REGION Network 10: Ethernet.Enc2 Too big speed change
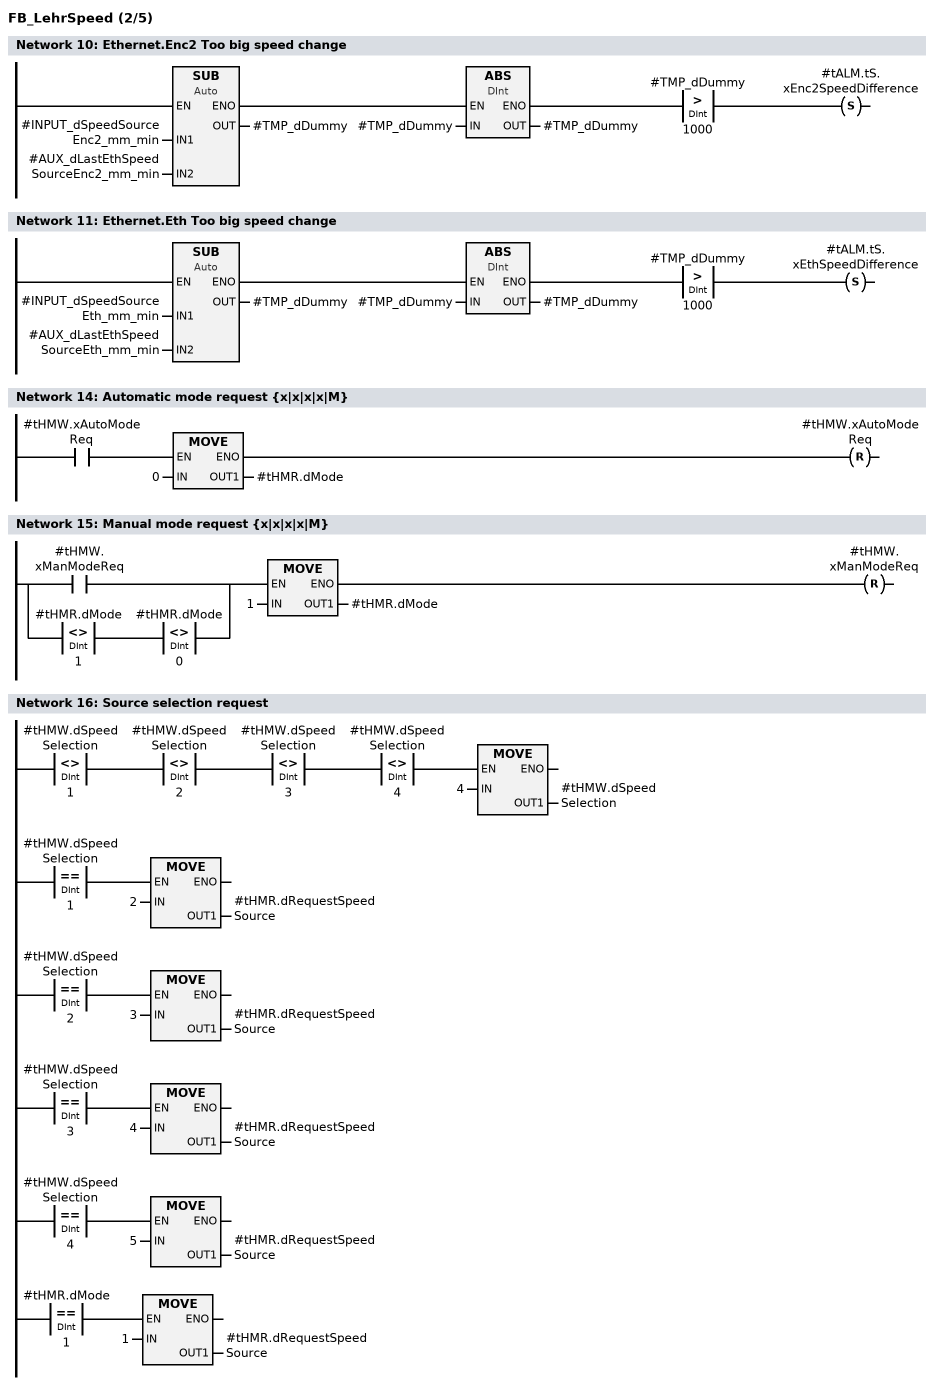
   RUNG wire#powerrail
      Sub(in1 := #INPUT_dSpeedSourceEnc2_mm_min, in2 := #AUX_dLastEthSpeedSourceEnc2_mm_min, out => #TMP_dDummy)
      { S7_Templates := "SrcType := DInt" } Abs(in := #TMP_dDummy, out => #TMP_dDummy)
      { S7_Templates := "SrcType := DInt" } GT_Contact(in1 := #TMP_dDummy, in2 := 1000)
      S_Coil( #tALM.tS.xEnc2SpeedDifference )
   END_RUNG
   // the same network as SCL:
   #TMP_dDummy := #INPUT_dSpeedSourceEnc2_mm_min - #AUX_dLastEthSpeedSourceEnc2_mm_min;
   #TMP_dDummy := ABS(#TMP_dDummy);
   IF #TMP_dDummy > 1000 THEN #tALM.tS.xEnc2SpeedDifference := TRUE; END_IF;
END_REGION

REGION Network 11: Ethernet.Eth Too big speed change
   RUNG wire#powerrail
      Sub(in1 := #INPUT_dSpeedSourceEth_mm_min, in2 := #AUX_dLastEthSpeedSourceEth_mm_min, out => #TMP_dDummy)
      { S7_Templates := "SrcType := DInt" } Abs(in := #TMP_dDummy, out => #TMP_dDummy)
      { S7_Templates := "SrcType := DInt" } GT_Contact(in1 := #TMP_dDummy, in2 := 1000)
      S_Coil( #tALM.tS.xEthSpeedDifference )
   END_RUNG
   // the same network as SCL:
   #TMP_dDummy := #INPUT_dSpeedSourceEth_mm_min - #AUX_dLastEthSpeedSourceEth_mm_min;
   #TMP_dDummy := ABS(#TMP_dDummy);
   IF #TMP_dDummy > 1000 THEN #tALM.tS.xEthSpeedDifference := TRUE; END_IF;
END_REGION

REGION Network 12 (SCL): Calculate cumulative statuses
       IF #tALM.tS.xEnc1OutOfRange OR #tALM.tS.xEnc1SpeedDifference THEN
           #ST_xStoppingFaultsEnc1 := TRUE;
       ELSE
           #ST_xStoppingFaultsEnc1 := FALSE;
       END_IF;

       IF #tALM.tS.xEnc2OutOfRange OR #tALM.tS.xEnc2SpeedDifference THEN
           #ST_xStoppingFaultsEnc2 := TRUE;
       ELSE
           #ST_xStoppingFaultsEnc2 := FALSE;
       END_IF;

       IF #tALM.tS.xEthOutOfRange OR #tALM.tS.xEthSpeedDifference OR #tALM.tS.xEthCommunicationTimeout THEN
           #ST_xStoppingFaultsEth := TRUE;
       ELSE
           #ST_xStoppingFaultsEth := FALSE;
       END_IF;

       GATHER(IN := #tALM.tF,
              OUT => #TMP_dwValue);

       IF #TMP_dwValue <> 0 THEN
           #ST_xFaults := TRUE;
       ELSE
           #ST_xFaults := FALSE;
       END_IF;

       GATHER(IN := #tALM.tW,
              OUT => #TMP_dwValue);

       IF #TMP_dwValue <> 0 THEN
           #ST_xWarnings := TRUE;
       ELSE
           #ST_xWarnings := FALSE;
       END_IF;
END_REGION

REGION Network 13: ####_HMI LOGICS_####
END_REGION

REGION Network 14: Automatic mode request {x|x|x|x|M}
   RUNG wire#powerrail
      Contact( #tHMW.xAutoModeReq )
      Move(in := 0, out1 => #tHMR.dMode)
      R_Coil( #tHMW.xAutoModeReq )
   END_RUNG
   // the same network as SCL:
   IF #tHMW.xAutoModeReq THEN
       #tHMR.dMode := 0;
       #tHMW.xAutoModeReq := FALSE;
   END_IF;
END_REGION

REGION Network 15: Manual mode request {x|x|x|x|M}
   RUNG wire#powerrail
      Contact( #tHMW.xManModeReq )
      wire#w1
      Move(in := 1, out1 => #tHMR.dMode)
      R_Coil( #tHMW.xManModeReq )
   END_RUNG
   RUNG wire#powerrail
      { S7_Templates := "SrcType := DInt" } NE_Contact(in1 := #tHMR.dMode, in2 := 1)
      { S7_Templates := "SrcType := DInt" } NE_Contact(in1 := #tHMR.dMode, in2 := 0)
   END_RUNG wire#w1
   // the same network as SCL:
   #_w1 := #tHMW.xManModeReq OR ((#tHMR.dMode <> 1) AND (#tHMR.dMode <> 0));
   IF #_w1 THEN
       #tHMR.dMode := 1;
       #tHMW.xManModeReq := FALSE;
   END_IF;
END_REGION

REGION Network 16: Source selection request
   RUNG wire#powerrail
      { S7_Templates := "SrcType := DInt" } NE_Contact(in1 := #tHMW.dSpeedSelection, in2 := 1)
      { S7_Templates := "SrcType := DInt" } NE_Contact(in1 := #tHMW.dSpeedSelection, in2 := 2)
      { S7_Templates := "SrcType := DInt" } NE_Contact(in1 := #tHMW.dSpeedSelection, in2 := 3)
      { S7_Templates := "SrcType := DInt" } NE_Contact(in1 := #tHMW.dSpeedSelection, in2 := 4)
      Move(in := 4, out1 => #tHMW.dSpeedSelection)
   END_RUNG
   RUNG wire#powerrail
      { S7_Templates := "SrcType := DInt" } EQ_Contact(in1 := #tHMW.dSpeedSelection, in2 := 1)
      Move(in := 2, out1 => #tHMR.dRequestSpeedSource)
   END_RUNG
   RUNG wire#powerrail
      { S7_Templates := "SrcType := DInt" } EQ_Contact(in1 := #tHMW.dSpeedSelection, in2 := 2)
      Move(in := 3, out1 => #tHMR.dRequestSpeedSource)
   END_RUNG
   RUNG wire#powerrail
      { S7_Templates := "SrcType := DInt" } EQ_Contact(in1 := #tHMW.dSpeedSelection, in2 := 3)
      Move(in := 4, out1 => #tHMR.dRequestSpeedSource)
   END_RUNG
   RUNG wire#powerrail
      { S7_Templates := "SrcType := DInt" } EQ_Contact(in1 := #tHMW.dSpeedSelection, in2 := 4)
      Move(in := 5, out1 => #tHMR.dRequestSpeedSource)
   END_RUNG
   RUNG wire#powerrail
      { S7_Templates := "SrcType := DInt" } EQ_Contact(in1 := #tHMR.dMode, in2 := 1)
      Move(in := 1, out1 => #tHMR.dRequestSpeedSource)
   END_RUNG
   // the same network as SCL:
   IF (#tHMW.dSpeedSelection <> 1) AND (#tHMW.dSpeedSelection <> 2) AND (#tHMW.dSpeedSelection <> 3) AND (#tHMW.dSpeedSelection <> 4) THEN
       #tHMW.dSpeedSelection := 4;
   END_IF;
   IF #tHMW.dSpeedSelection = 1 THEN #tHMR.dRequestSpeedSource := 2; END_IF;
   IF #tHMW.dSpeedSelection = 2 THEN #tHMR.dRequestSpeedSource := 3; END_IF;
   IF #tHMW.dSpeedSelection = 3 THEN #tHMR.dRequestSpeedSource := 4; END_IF;
   IF #tHMW.dSpeedSelection = 4 THEN #tHMR.dRequestSpeedSource := 5; END_IF;
   IF #tHMR.dMode = 1 THEN #tHMR.dRequestSpeedSource := 1; END_IF;
END_REGION

REGION Network 17: ###_STATUSES_###
END_REGION

REGION Network 18: Update speeds
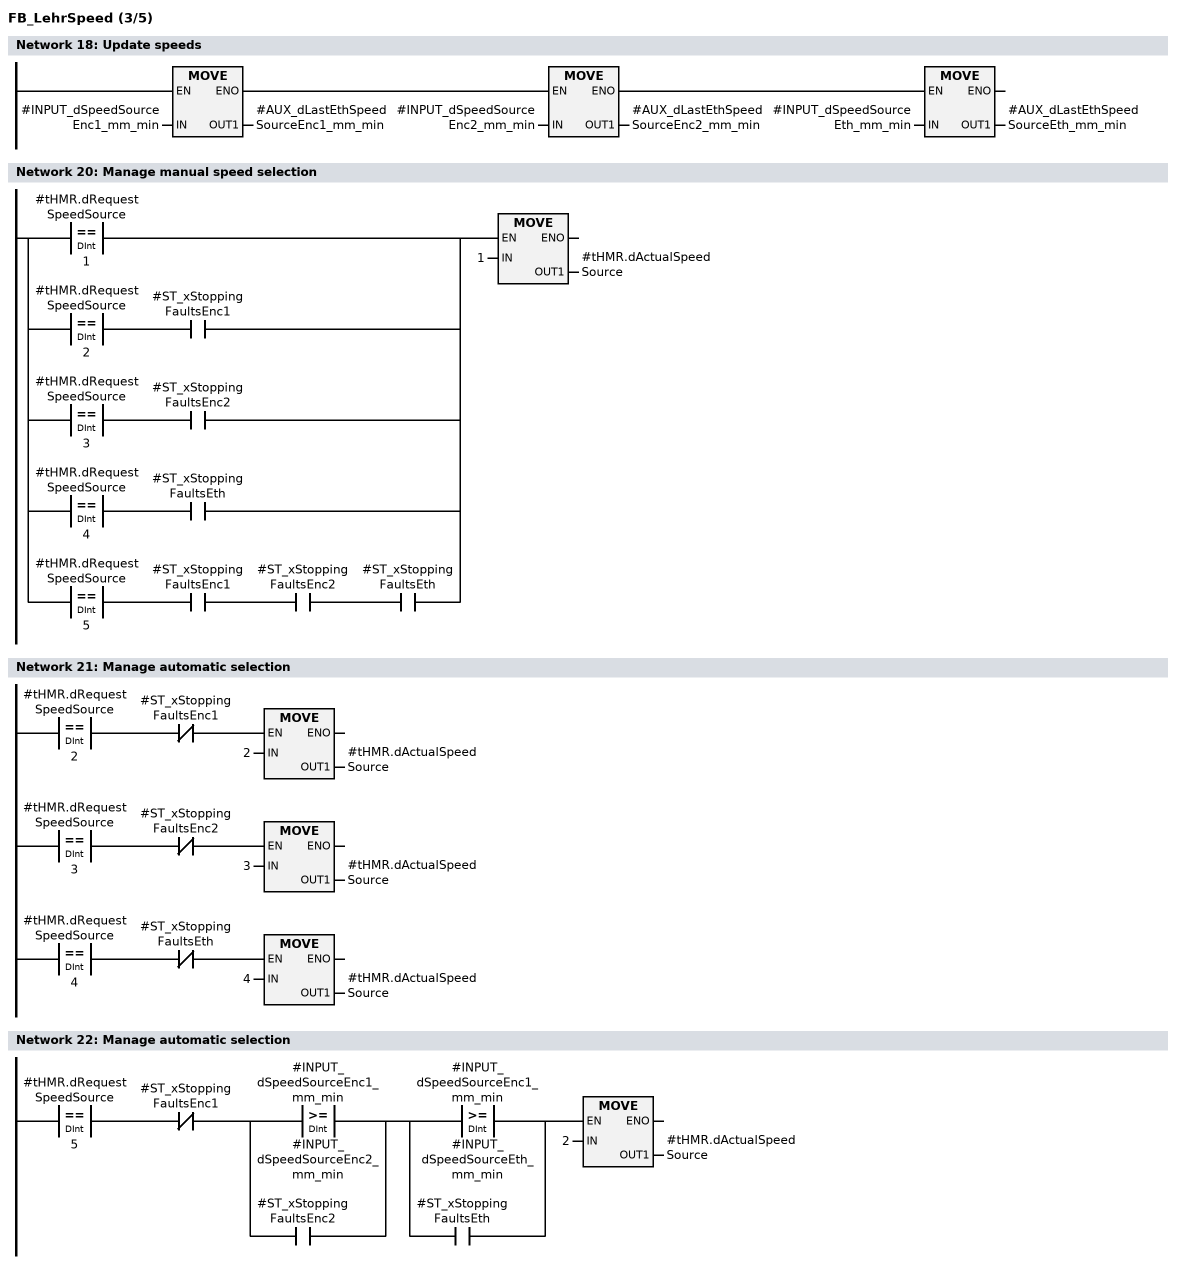
   RUNG wire#powerrail
      Move(in := #INPUT_dSpeedSourceEnc1_mm_min, out1 => #AUX_dLastEthSpeedSourceEnc1_mm_min)
      Move(in := #INPUT_dSpeedSourceEnc2_mm_min, out1 => #AUX_dLastEthSpeedSourceEnc2_mm_min)
      Move(in := #INPUT_dSpeedSourceEth_mm_min, out1 => #AUX_dLastEthSpeedSourceEth_mm_min)
   END_RUNG
   // the same network as SCL:
   #AUX_dLastEthSpeedSourceEnc1_mm_min := #INPUT_dSpeedSourceEnc1_mm_min;
   #AUX_dLastEthSpeedSourceEnc2_mm_min := #INPUT_dSpeedSourceEnc2_mm_min;
   #AUX_dLastEthSpeedSourceEth_mm_min := #INPUT_dSpeedSourceEth_mm_min;
END_REGION

REGION Network 19: ###_PHASES_&_LOGICS_###
END_REGION

REGION Network 20: Manage manual speed selection
   RUNG wire#powerrail
      { S7_Templates := "SrcType := DInt" } EQ_Contact(in1 := #tHMR.dRequestSpeedSource, in2 := 1)
      wire#w1
      Move(in := 1, out1 => #tHMR.dActualSpeedSource)
   END_RUNG
   RUNG wire#powerrail
      { S7_Templates := "SrcType := DInt" } EQ_Contact(in1 := #tHMR.dRequestSpeedSource, in2 := 2)
      Contact( #ST_xStoppingFaultsEnc1 )
   END_RUNG wire#w1
   RUNG wire#powerrail
      { S7_Templates := "SrcType := DInt" } EQ_Contact(in1 := #tHMR.dRequestSpeedSource, in2 := 3)
      Contact( #ST_xStoppingFaultsEnc2 )
   END_RUNG wire#w1
   RUNG wire#powerrail
      { S7_Templates := "SrcType := DInt" } EQ_Contact(in1 := #tHMR.dRequestSpeedSource, in2 := 4)
      Contact( #ST_xStoppingFaultsEth )
   END_RUNG wire#w1
   RUNG wire#powerrail
      { S7_Templates := "SrcType := DInt" } EQ_Contact(in1 := #tHMR.dRequestSpeedSource, in2 := 5)
      Contact( #ST_xStoppingFaultsEnc1 )
      Contact( #ST_xStoppingFaultsEnc2 )
      Contact( #ST_xStoppingFaultsEth )
   END_RUNG wire#w1
   // the same network as SCL:
   IF (#tHMR.dRequestSpeedSource = 1) OR ((#tHMR.dRequestSpeedSource = 2) AND #ST_xStoppingFaultsEnc1) OR ((#tHMR.dRequestSpeedSource = 3) AND #ST_xStoppingFaultsEnc2) OR ((#tHMR.dRequestSpeedSource = 4) AND #ST_xStoppingFaultsEth) OR ((#tHMR.dRequestSpeedSource = 5) AND #ST_xStoppingFaultsEnc1 AND #ST_xStoppingFaultsEnc2 AND #ST_xStoppingFaultsEth) THEN
       #tHMR.dActualSpeedSource := 1;
   END_IF;
END_REGION

REGION Network 21: Manage automatic selection
   RUNG wire#powerrail
      { S7_Templates := "SrcType := DInt" } EQ_Contact(in1 := #tHMR.dRequestSpeedSource, in2 := 2)
      I_Contact( #ST_xStoppingFaultsEnc1 )
      Move(in := 2, out1 => #tHMR.dActualSpeedSource)
   END_RUNG
   RUNG wire#powerrail
      { S7_Templates := "SrcType := DInt" } EQ_Contact(in1 := #tHMR.dRequestSpeedSource, in2 := 3)
      I_Contact( #ST_xStoppingFaultsEnc2 )
      Move(in := 3, out1 => #tHMR.dActualSpeedSource)
   END_RUNG
   RUNG wire#powerrail
      { S7_Templates := "SrcType := DInt" } EQ_Contact(in1 := #tHMR.dRequestSpeedSource, in2 := 4)
      I_Contact( #ST_xStoppingFaultsEth )
      Move(in := 4, out1 => #tHMR.dActualSpeedSource)
   END_RUNG
   // the same network as SCL:
   IF (#tHMR.dRequestSpeedSource = 2) AND NOT #ST_xStoppingFaultsEnc1 THEN
       #tHMR.dActualSpeedSource := 2;
   END_IF;
   IF (#tHMR.dRequestSpeedSource = 3) AND NOT #ST_xStoppingFaultsEnc2 THEN
       #tHMR.dActualSpeedSource := 3;
   END_IF;
   IF (#tHMR.dRequestSpeedSource = 4) AND NOT #ST_xStoppingFaultsEth THEN
       #tHMR.dActualSpeedSource := 4;
   END_IF;
END_REGION

REGION Network 22: Manage automatic selection
   RUNG wire#powerrail
      { S7_Templates := "SrcType := DInt" } EQ_Contact(in1 := #tHMR.dRequestSpeedSource, in2 := 5)
      I_Contact( #ST_xStoppingFaultsEnc1 )
      wire#w1
      { S7_Templates := "SrcType := DInt" } GE_Contact(in1 := #INPUT_dSpeedSourceEnc1_mm_min, in2 := #INPUT_dSpeedSourceEnc2_mm_min)
      wire#w2
      { S7_Templates := "SrcType := DInt" } GE_Contact(in1 := #INPUT_dSpeedSourceEnc1_mm_min, in2 := #INPUT_dSpeedSourceEth_mm_min)
      wire#w3
      Move(in := 2, out1 => #tHMR.dActualSpeedSource)
   END_RUNG
   RUNG wire#w1
      Contact( #ST_xStoppingFaultsEnc2 )
   END_RUNG wire#w2
   RUNG wire#w2
      Contact( #ST_xStoppingFaultsEth )
   END_RUNG wire#w3
   // the same network as SCL:
   IF (#tHMR.dRequestSpeedSource = 5) AND NOT #ST_xStoppingFaultsEnc1 AND ((#INPUT_dSpeedSourceEnc1_mm_min >= #INPUT_dSpeedSourceEnc2_mm_min) OR #ST_xStoppingFaultsEnc2) AND ((#INPUT_dSpeedSourceEnc1_mm_min >= #INPUT_dSpeedSourceEth_mm_min) OR #ST_xStoppingFaultsEth) THEN
       #tHMR.dActualSpeedSource := 2;
   END_IF;
END_REGION

REGION Network 23: Manage automatic selection
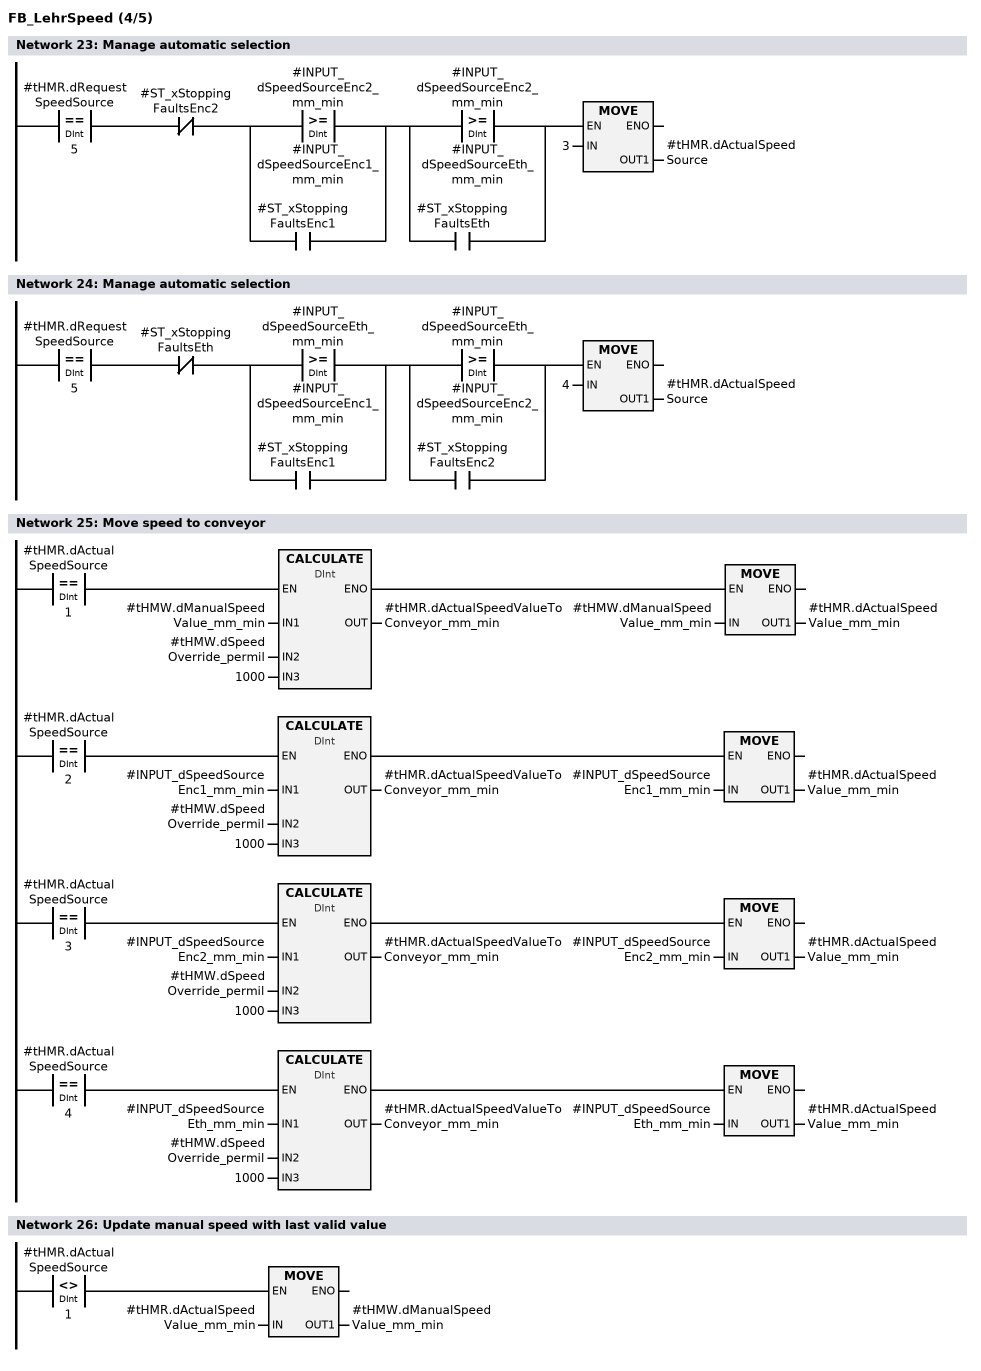
   RUNG wire#powerrail
      { S7_Templates := "SrcType := DInt" } EQ_Contact(in1 := #tHMR.dRequestSpeedSource, in2 := 5)
      I_Contact( #ST_xStoppingFaultsEnc2 )
      wire#w1
      { S7_Templates := "SrcType := DInt" } GE_Contact(in1 := #INPUT_dSpeedSourceEnc2_mm_min, in2 := #INPUT_dSpeedSourceEnc1_mm_min)
      wire#w2
      { S7_Templates := "SrcType := DInt" } GE_Contact(in1 := #INPUT_dSpeedSourceEnc2_mm_min, in2 := #INPUT_dSpeedSourceEth_mm_min)
      wire#w3
      Move(in := 3, out1 => #tHMR.dActualSpeedSource)
   END_RUNG
   RUNG wire#w1
      Contact( #ST_xStoppingFaultsEnc1 )
   END_RUNG wire#w2
   RUNG wire#w2
      Contact( #ST_xStoppingFaultsEth )
   END_RUNG wire#w3
   // the same network as SCL:
   IF (#tHMR.dRequestSpeedSource = 5) AND NOT #ST_xStoppingFaultsEnc2 AND ((#INPUT_dSpeedSourceEnc2_mm_min >= #INPUT_dSpeedSourceEnc1_mm_min) OR #ST_xStoppingFaultsEnc1) AND ((#INPUT_dSpeedSourceEnc2_mm_min >= #INPUT_dSpeedSourceEth_mm_min) OR #ST_xStoppingFaultsEth) THEN
       #tHMR.dActualSpeedSource := 3;
   END_IF;
END_REGION

REGION Network 24: Manage automatic selection
   RUNG wire#powerrail
      { S7_Templates := "SrcType := DInt" } EQ_Contact(in1 := #tHMR.dRequestSpeedSource, in2 := 5)
      I_Contact( #ST_xStoppingFaultsEth )
      wire#w1
      { S7_Templates := "SrcType := DInt" } GE_Contact(in1 := #INPUT_dSpeedSourceEth_mm_min, in2 := #INPUT_dSpeedSourceEnc1_mm_min)
      wire#w2
      { S7_Templates := "SrcType := DInt" } GE_Contact(in1 := #INPUT_dSpeedSourceEth_mm_min, in2 := #INPUT_dSpeedSourceEnc2_mm_min)
      wire#w3
      Move(in := 4, out1 => #tHMR.dActualSpeedSource)
   END_RUNG
   RUNG wire#w1
      Contact( #ST_xStoppingFaultsEnc1 )
   END_RUNG wire#w2
   RUNG wire#w2
      Contact( #ST_xStoppingFaultsEnc2 )
   END_RUNG wire#w3
   // the same network as SCL:
   IF (#tHMR.dRequestSpeedSource = 5) AND NOT #ST_xStoppingFaultsEth AND ((#INPUT_dSpeedSourceEth_mm_min >= #INPUT_dSpeedSourceEnc1_mm_min) OR #ST_xStoppingFaultsEnc1) AND ((#INPUT_dSpeedSourceEth_mm_min >= #INPUT_dSpeedSourceEnc2_mm_min) OR #ST_xStoppingFaultsEnc2) THEN
       #tHMR.dActualSpeedSource := 4;
   END_IF;
END_REGION

REGION Network 25: Move speed to conveyor
   RUNG wire#powerrail
      { S7_Templates := "SrcType := DInt" } EQ_Contact(in1 := #tHMR.dActualSpeedSource, in2 := 1)
      { S7_Templates := "SrcType := DInt"; S7_Expression := "IN1+(IN1/IN3*IN2)" } Calculate(in1 := #tHMW.dManualSpeedValue_mm_min, in2 := #tHMW.dSpeedOverride_permil, in3 := 1000, out => #tHMR.dActualSpeedValueToConveyor_mm_min)
      Move(in := #tHMW.dManualSpeedValue_mm_min, out1 => #tHMR.dActualSpeedValue_mm_min)
   END_RUNG
   RUNG wire#powerrail
      { S7_Templates := "SrcType := DInt" } EQ_Contact(in1 := #tHMR.dActualSpeedSource, in2 := 2)
      { S7_Templates := "SrcType := DInt"; S7_Expression := "IN1+(IN1/IN3*IN2)" } Calculate(in1 := #INPUT_dSpeedSourceEnc1_mm_min, in2 := #tHMW.dSpeedOverride_permil, in3 := 1000, out => #tHMR.dActualSpeedValueToConveyor_mm_min)
      Move(in := #INPUT_dSpeedSourceEnc1_mm_min, out1 => #tHMR.dActualSpeedValue_mm_min)
   END_RUNG
   RUNG wire#powerrail
      { S7_Templates := "SrcType := DInt" } EQ_Contact(in1 := #tHMR.dActualSpeedSource, in2 := 3)
      { S7_Templates := "SrcType := DInt"; S7_Expression := "IN1+(IN1/IN3*IN2)" } Calculate(in1 := #INPUT_dSpeedSourceEnc2_mm_min, in2 := #tHMW.dSpeedOverride_permil, in3 := 1000, out => #tHMR.dActualSpeedValueToConveyor_mm_min)
      Move(in := #INPUT_dSpeedSourceEnc2_mm_min, out1 => #tHMR.dActualSpeedValue_mm_min)
   END_RUNG
   RUNG wire#powerrail
      { S7_Templates := "SrcType := DInt" } EQ_Contact(in1 := #tHMR.dActualSpeedSource, in2 := 4)
      { S7_Templates := "SrcType := DInt"; S7_Expression := "IN1+(IN1/IN3*IN2)" } Calculate(in1 := #INPUT_dSpeedSourceEth_mm_min, in2 := #tHMW.dSpeedOverride_permil, in3 := 1000, out => #tHMR.dActualSpeedValueToConveyor_mm_min)
      Move(in := #INPUT_dSpeedSourceEth_mm_min, out1 => #tHMR.dActualSpeedValue_mm_min)
   END_RUNG
   // the same network as SCL:
   IF #tHMR.dActualSpeedSource = 1 THEN
       #tHMR.dActualSpeedValueToConveyor_mm_min := #tHMW.dManualSpeedValue_mm_min+(#tHMW.dManualSpeedValue_mm_min/1000*#tHMW.dSpeedOverride_permil);
       #tHMR.dActualSpeedValue_mm_min := #tHMW.dManualSpeedValue_mm_min;
   END_IF;
   IF #tHMR.dActualSpeedSource = 2 THEN
       #tHMR.dActualSpeedValueToConveyor_mm_min := #INPUT_dSpeedSourceEnc1_mm_min+(#INPUT_dSpeedSourceEnc1_mm_min/1000*#tHMW.dSpeedOverride_permil);
       #tHMR.dActualSpeedValue_mm_min := #INPUT_dSpeedSourceEnc1_mm_min;
   END_IF;
   IF #tHMR.dActualSpeedSource = 3 THEN
       #tHMR.dActualSpeedValueToConveyor_mm_min := #INPUT_dSpeedSourceEnc2_mm_min+(#INPUT_dSpeedSourceEnc2_mm_min/1000*#tHMW.dSpeedOverride_permil);
       #tHMR.dActualSpeedValue_mm_min := #INPUT_dSpeedSourceEnc2_mm_min;
   END_IF;
   IF #tHMR.dActualSpeedSource = 4 THEN
       #tHMR.dActualSpeedValueToConveyor_mm_min := #INPUT_dSpeedSourceEth_mm_min+(#INPUT_dSpeedSourceEth_mm_min/1000*#tHMW.dSpeedOverride_permil);
       #tHMR.dActualSpeedValue_mm_min := #INPUT_dSpeedSourceEth_mm_min;
   END_IF;
END_REGION

REGION Network 26: Update manual speed with last valid value
   RUNG wire#powerrail
      { S7_Templates := "SrcType := DInt" } NE_Contact(in1 := #tHMR.dActualSpeedSource, in2 := 1)
      Move(in := #tHMR.dActualSpeedValue_mm_min, out1 => #tHMW.dManualSpeedValue_mm_min)
   END_RUNG
   // the same network as SCL:
   IF #tHMR.dActualSpeedSource <> 1 THEN
       #tHMW.dManualSpeedValue_mm_min := #tHMR.dActualSpeedValue_mm_min;
   END_IF;
END_REGION

REGION Network 27: ###_HMI_STATUSES_###
END_REGION

REGION Network 28: Status hmi
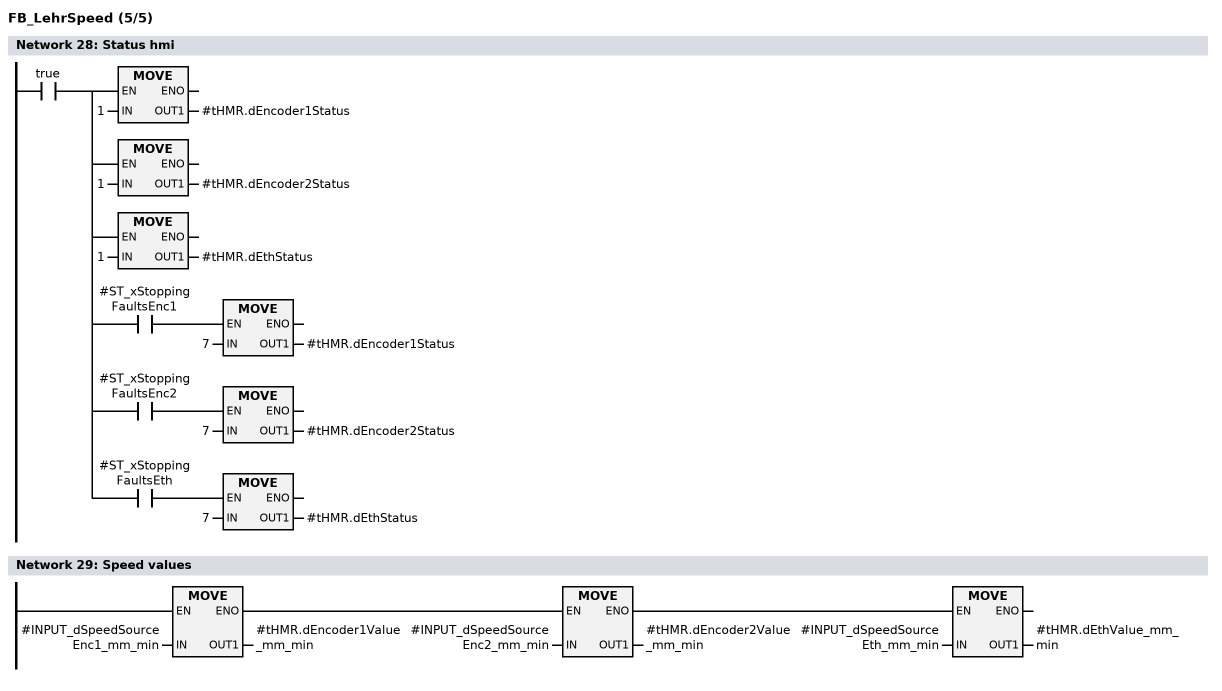
   RUNG wire#powerrail
      Contact( true )
      wire#w1
      Move(in := 1, out1 => #tHMR.dEncoder1Status)
   END_RUNG
   RUNG wire#w1
      Move(in := 1, out1 => #tHMR.dEncoder2Status)
   END_RUNG
   RUNG wire#w1
      Move(in := 1, out1 => #tHMR.dEthStatus)
   END_RUNG
   RUNG wire#w1
      Contact( #ST_xStoppingFaultsEnc1 )
      Move(in := 7, out1 => #tHMR.dEncoder1Status)
   END_RUNG
   RUNG wire#w1
      Contact( #ST_xStoppingFaultsEnc2 )
      Move(in := 7, out1 => #tHMR.dEncoder2Status)
   END_RUNG
   RUNG wire#w1
      Contact( #ST_xStoppingFaultsEth )
      Move(in := 7, out1 => #tHMR.dEthStatus)
   END_RUNG
   // the same network as SCL:
   IF true THEN
       #tHMR.dEncoder1Status := 1;
       #tHMR.dEncoder2Status := 1;
       #tHMR.dEthStatus := 1;
   END_IF;
   IF true AND #ST_xStoppingFaultsEnc1 THEN #tHMR.dEncoder1Status := 7; END_IF;
   IF true AND #ST_xStoppingFaultsEnc2 THEN #tHMR.dEncoder2Status := 7; END_IF;
   IF true AND #ST_xStoppingFaultsEth THEN #tHMR.dEthStatus := 7; END_IF;
END_REGION

REGION Network 29: Speed values
   RUNG wire#powerrail
      Move(in := #INPUT_dSpeedSourceEnc1_mm_min, out1 => #tHMR.dEncoder1Value_mm_min)
      Move(in := #INPUT_dSpeedSourceEnc2_mm_min, out1 => #tHMR.dEncoder2Value_mm_min)
      Move(in := #INPUT_dSpeedSourceEth_mm_min, out1 => #tHMR.dEthValue_mm_min)
   END_RUNG
   // the same network as SCL:
   #tHMR.dEncoder1Value_mm_min := #INPUT_dSpeedSourceEnc1_mm_min;
   #tHMR.dEncoder2Value_mm_min := #INPUT_dSpeedSourceEnc2_mm_min;
   #tHMR.dEthValue_mm_min := #INPUT_dSpeedSourceEth_mm_min;
END_REGION

REGION Network 30 (SCL): Lehr position advancement [mm/100]
   #AUX_dLehrPositionAdvancement := (REAL_TO_DINT(DINT_TO_REAL(#tHMR.dActualSpeedValue_mm_min * 100) / 60000.0) * "GP_OB_Initialize_Slow_IDB".OUT_dExecutionTime_ms) + #AUX_dLehrPositionAdvancement;
END_REGION
END_FUNCTION_BLOCK

FUNCTION "Z200_SpeedLehr" : Void   // FC112, LAD
{ S7_Optimized_Access := 'TRUE' }
VERSION : 0.1
   VAR_TEMP
      TMP_xGetPulseEncoder : Bool;
      TMP_dDifferenceMeasureEnc1 : DInt;
      TMP_dDifferenceMeasureEnc2 : DInt;
      TMP_d : DInt;
   END_VAR
   VAR CONSTANT
      CONST_rKConvEnc1 : Real := 17.8729;
      CONST_rKConvEnc2 : Real := 17.8729;
   END_VAR
BEGIN

REGION Network 1
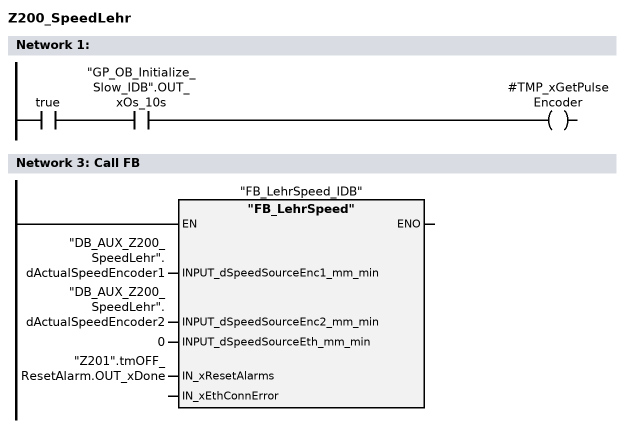
   RUNG wire#powerrail
      Contact( true )
      Contact( "GP_OB_Initialize_Slow_IDB".OUT_xOs_10s )
      Coil( #TMP_xGetPulseEncoder )
   END_RUNG
   // the same network as SCL:
   #TMP_xGetPulseEncoder := true AND "GP_OB_Initialize_Slow_IDB".OUT_xOs_10s;
END_REGION

REGION Network 2 (SCL): Encoder Speed Calculation
   IF #TMP_xGetPulseEncoder THEN
       #TMP_dDifferenceMeasureEnc1 := "DB_AUX_Z200_SpeedLehr".dPulseEncoder1 - "DB_AUX_Z200_SpeedLehr".dLastPulseEnc1;
       #TMP_dDifferenceMeasureEnc2 := "DB_AUX_Z200_SpeedLehr".dPulseEncoder2 - "DB_AUX_Z200_SpeedLehr".dLastPulseEnc2;
       //Enc 1


       IF #TMP_dDifferenceMeasureEnc1 > 0 THEN

           "DB_AUX_Z200_SpeedLehr".dActualSpeedEncoder1 := REAL_TO_DINT(DINT_TO_REAL(#TMP_dDifferenceMeasureEnc1) / #CONST_rKConvEnc1);
           "DB_AUX_Z200_SpeedLehr".dActualSpeedEncoder2 := REAL_TO_DINT(DINT_TO_REAL(#TMP_dDifferenceMeasureEnc2) / #CONST_rKConvEnc1);

       END_IF;

       "DB_AUX_Z200_SpeedLehr".dLastPulseEnc1 := "DB_AUX_Z200_SpeedLehr".dPulseEncoder1;
       "DB_AUX_Z200_SpeedLehr".dLastPulseEnc2 := "DB_AUX_Z200_SpeedLehr".dPulseEncoder2;

   END_IF;
END_REGION

REGION Network 3: Call FB
   RUNG wire#powerrail
      "FB_LehrSpeed_IDB"(INPUT_dSpeedSourceEnc1_mm_min := "DB_AUX_Z200_SpeedLehr".dActualSpeedEncoder1, INPUT_dSpeedSourceEnc2_mm_min := "DB_AUX_Z200_SpeedLehr".dActualSpeedEncoder2, INPUT_dSpeedSourceEth_mm_min := 0, IN_xResetAlarms := "Z201".tmOFF_ResetAlarm.OUT_xDone, IN_xEthConnError :=)
   END_RUNG
   // the same network as SCL:
   "FB_LehrSpeed_IDB"(INPUT_dSpeedSourceEnc1_mm_min := "DB_AUX_Z200_SpeedLehr".dActualSpeedEncoder1,   // "FB_LehrSpeed"
                      INPUT_dSpeedSourceEnc2_mm_min := "DB_AUX_Z200_SpeedLehr".dActualSpeedEncoder2,
                      INPUT_dSpeedSourceEth_mm_min := 0,
                      IN_xResetAlarms := "Z201".tmOFF_ResetAlarm.OUT_xDone);
END_REGION
END_FUNCTION

// folder: 03_Programs_Logics/MCC1201/29_Sinamics

FUNCTION_BLOCK "SINAMICS_ControlUnit"   // FB50, LAD
{ S7_Optimized_Access := 'FALSE' }
AUTHOR : Armitano
VERSION : 1.7
// Return value:
// * 0: OK
// Blocking message:
// * group 1 to 9: general error
// * group 10 to 19: system data error
//   * 10: Sinamics input/output addresses for control unit wrong or not setted
//   * 11: Sinamics input/output addresses for power module wrong 
//   * 12: Delay time before shut down too low or not setted
   VAR_INPUT
      IN_xSwitching_EN : Bool;   // Switching on for power module
      IN_xResetFaults : Bool;   // Reset faults
   END_VAR
   VAR_OUTPUT
      OUT_xPower_ON : Bool;   // Power module switched on
      OUT_xCU_FaultPresent : Bool;   // Control unit fault present
      OUT_xPM_FaultPresent : Bool;   // Power module fault present
      OUT_xRetVal : Int;   // Return value in case of wrong configuration
   END_VAR
   VAR
      STC_tSYS_DATA : Struct   // System data
         iIOAddress_CU : Int := -1;   // Input/Output addresses for control unit
         iIOAddress_PM : Int := -1;   // Input/Output addresses for power module [0=No power module]
         iPowerOFFDelay_ms : Int := 1000;   // Delay time before shut down [ms]
      END_STRUCT;
      STC_tPH : Struct
         x0 : Bool;   // Shut down delay
         x1 : Bool;   // Power ON delay
         x2 : Bool;
         x3 : Bool;
         x4 : Bool;
         x5 : Bool;
         x6 : Bool;
         x7 : Bool;
         x8 : Bool;
         x9 : Bool;
         x10 : Bool;
         x11 : Bool;
         x12 : Bool;
         x13 : Bool;
         x14 : Bool;
         x15 : Bool;
      END_STRUCT;
      STC_tPROP : Struct
         i0 : Int;   // Previous cycle [ms]
         tmOFF_DelayOFF_ms : IEC_TIMER;   // Delay shut down [ms]
         tmON_DelayON_ms : IEC_TIMER;   // Delay power ON [ms]
         i3 : Int;
         i4 : Int;
      END_STRUCT;
      STC_tPZD_CU : Struct   // Control unit telegram
         tR : Struct   // READ
            tZSW1 : Struct   // R2089[1].STATUS WORD 1
               x8 : Bool;   // System time synchronized
               x9 : Bool;   // Group alarm present
               x10 : Bool;   // Group fault present
               x11 : Bool;   // Safety group message present
               x12 : Bool;   // Slave sign of life bit 0
               x13 : Bool;   // Slave sign of life bit 1
               x14 : Bool;   // Slave sign of life bit 2
               x15 : Bool;   // Slave sign of life bit 3
               x0 : Bool;   // Reserved
               x1 : Bool;   // Reserved
               x2 : Bool;   // Reserved
               x3 : Bool;   // Fault present
               x4 : Bool;   // Reserved
               x5 : Bool;   // Reserved
               x6 : Bool;   // Reserved
               x7 : Bool;   // Alarm present
            END_STRUCT;
            tE_DIGITAL : Struct   // R2089[2].DIGITAL INPUT WORD 1
               x8 : Bool;   // DI 0
               x9 : Bool;   // DI 1
               x10 : Bool;   // DI 2
               x11 : Bool;   // DI 3
               x12 : Bool;   // DI 4
               x13 : Bool;   // DI 5
               x14 : Bool;   // DI 6
               x15 : Bool;   // DI 7
               x0 : Bool;   // DI/DO 8
               x1 : Bool;   // DI/DO 9
               x2 : Bool;   // DI/DO 10
               x3 : Bool;   // DI/DO 11
               x4 : Bool;   // DI/DO 12
               x5 : Bool;   // DI/DO 13
               x6 : Bool;   // DI/DO 14
               x7 : Bool;   // DI/DO 15
            END_STRUCT;
            tE_DIGITAL_1 : Struct   // R2089[3].DIGITAL INPUT WORD 2
               x8 : Bool;   // DI 16
               x9 : Bool;   // DI 17
               x10 : Bool;   // Reserved
               x11 : Bool;   // Reserved
               x12 : Bool;   // DI 20
               x13 : Bool;   // DI 21
               x14 : Bool;   // Reserved
               x15 : Bool;   // Reserved
               x0 : Bool;   // Reserved
               x1 : Bool;   // Reserved
               x2 : Bool;   // Reserved
               x3 : Bool;   // Reserved
               x4 : Bool;   // Reserved
               x5 : Bool;   // Reserved
               x6 : Bool;   // Reserved
               x7 : Bool;   // Reserved
            END_STRUCT;
         END_STRUCT;
         tW : Struct   // WRITE
            tSTW1 : Struct   // CONTROL WORD 1
               x8 : Bool;   // Reserved
               x9 : Bool;   // Reserved
               x10 : Bool;   // P3116.Acknowledgment automatically suppressed
               x11 : Bool;   // Reserved
               x12 : Bool;   // Master sign of life bit0
               x13 : Bool;   // Master sign of life bit1
               x14 : Bool;   // Master sign of life bit2
               x15 : Bool;   // Master sign of life bit3
               x0 : Bool;   // P681.Central misuring probe, synchronizing signal source
               x1 : Bool;   // P3104.RTC real time synchronization PING
               x2 : Bool;   // Reserved
               x3 : Bool;   // Reserved
               x4 : Bool;   // Reserved
               x5 : Bool;   // Reserved
               x6 : Bool;   // Reserved
               x7 : Bool;   // P2103.Acknowledgment faults
            END_STRUCT;
            tA_DIGITAL : Struct   // DIGITAL OUTPUT WORD 1
               x8 : Bool;   // Reserved
               x9 : Bool;   // Reserved
               x10 : Bool;   // Reserved
               x11 : Bool;   // Reserved
               x12 : Bool;   // Reserved
               x13 : Bool;   // Reserved
               x14 : Bool;   // Reserved
               x15 : Bool;   // Reserved
               x0 : Bool;   // P738.CU, signal source for terminal DI/DO 8
               x1 : Bool;   // P739.CU, signal source for terminal DI/DO 9
               x2 : Bool;   // P740.CU, signal source for terminal DI/DO 10
               x3 : Bool;   // P741.CU, signal source for terminal DI/DO 11
               x4 : Bool;   // P742.CU, signal source for terminal DI/DO 12
               x5 : Bool;   // P743.CU, signal source for terminal DI/DO 13
               x6 : Bool;   // P744.CU, signal source for terminal DI/DO 14
               x7 : Bool;   // P745.CU, signal source for terminal DI/DO 15
            END_STRUCT;
            tA_DIGITAL_1 : Struct   // DIGITAL OUTPUT WORD 2
               x8 : Bool;   // Reserved
               x9 : Bool;   // Reserved
               x10 : Bool;   // Reserved
               x11 : Bool;   // Reserved
               x12 : Bool;   // Reserved
               x13 : Bool;   // Reserved
               x14 : Bool;   // Reserved
               x15 : Bool;   // Reserved
               x0 : Bool;   // Reserved
               x1 : Bool;   // Reserved
               x2 : Bool;   // Reserved
               x3 : Bool;   // Reserved
               x4 : Bool;   // Reserved
               x5 : Bool;   // Reserved
               x6 : Bool;   // Reserved
               x7 : Bool;   // Reserved
            END_STRUCT;
         END_STRUCT;
      END_STRUCT;
      STC_tPZD_PM : Struct   // Power module telegram
         tR : Struct   // READ
            tZSW1 : Struct   // P2089[0].STATUS WORD 1
               x8 : Bool;   // Reserved
               x9 : Bool;   // Control request
               x10 : Bool;   // Reserved
               x11 : Bool;   // Pre-charging completed
               x12 : Bool;   // Line contactor closed
               x13 : Bool;   // Reserved
               x14 : Bool;   // Reserved
               x15 : Bool;   // Reserved
               x0 : Bool;   // Ready for switch ON
               x1 : Bool;   // Ready
               x2 : Bool;   // Operation enabled
               x3 : Bool;   // Fault present
               x4 : Bool;   // No OFF2 active
               x5 : Bool;   // Reserved
               x6 : Bool;   // Sw on inhibit
               x7 : Bool;   // Alarm present
            END_STRUCT;
         END_STRUCT;
         tW : Struct   // WRITE
            tSTW1 : Struct   // CONTROL WORD 1
               x8 : Bool;   // Reserved
               x9 : Bool;   // Reserved
               x10 : Bool;   // P854[0].Control by PLC
               x11 : Bool;   // Reserved
               x12 : Bool;   // Reserved
               x13 : Bool;   // Reserved
               x14 : Bool;   // Reserved
               x15 : Bool;   // Reserved
               x0 : Bool;   // P840[0].ON/OFF
               x1 : Bool;   // P844[0].OFF2
               x2 : Bool;   // Reserved
               x3 : Bool;   // P852[0].Enable operation
               x4 : Bool;   // Reserved
               x5 : Bool;   // P3532.Inhibit monitoring
               x6 : Bool;   // P3533.Inhibit generator mode
               x7 : Bool;   // P2103[0].Acknowledge faults
            END_STRUCT;
         END_STRUCT;
      END_STRUCT;
   END_VAR
   VAR_TEMP
      TMP_dOldValue_AR1 : DInt;
      TMP_dOldValue_AR2 : DInt;
      TMP_x : Bool;
      TMP_i : Int;
      TMP_d : DInt;
      TMP_r : Real;
      TMP_a : ANY;
      TMP_tm : Time;
      TMP_dZero : DInt;
      TMP_xAlwaysON : Bool;
      TMP_dIO_Pointer : DInt;
      TMP_dPZD_Pointer : DInt;
   END_VAR
BEGIN

REGION Network 1 (STL): Save AR1 & AR2 value
   //    TAR1
   //    T     #OldValue_AR1
   //    TAR2
   //    T     #OldValue_AR2
END_REGION

REGION Network 2: #####_COSTANTS_#####
END_REGION

REGION Network 3 (STL): Initializing
         SET;
         S     #TMP_xAlwaysON;

         L     0;
         T     #OUT_xRetVal;

         L     DINT#0;
         T     #TMP_dZero;

         CALL  FILL
         ( BVAL    := #TMP_dZero,
           RET_VAL := #OUT_xRetVal,
           BLK     := #STC_tPZD_CU.tR
         );

         CALL  FILL
         ( BVAL    := #TMP_dZero,
           RET_VAL := #OUT_xRetVal,
           BLK     := #STC_tPZD_PM.tR
         );
END_REGION

REGION Network 4: #####_MATCH_#####
END_REGION

REGION Network 5 (STL): Input copy control unit
         L     #STC_tSYS_DATA.iIOAddress_CU;
         L     0;
         <I;
         JC    NWPM;

         L     #STC_tSYS_DATA.iIOAddress_CU;
         SLW   3;
         T     #TMP_dIO_Pointer;

         L;
         T     #TMP_dPZD_Pointer;

         L     IW[ #TMP_dIO_Pointer];
         T     DIW[ #TMP_dPZD_Pointer];

         L     #TMP_dIO_Pointer;
         +     16;
         T     #TMP_dIO_Pointer;
         L     #TMP_dPZD_Pointer;
         +     16;
         T     #TMP_dPZD_Pointer;

         L     IW[ #TMP_dIO_Pointer];
         T     DIW[ #TMP_dPZD_Pointer];

         L     #TMP_dIO_Pointer;
         +     16;
         T     #TMP_dIO_Pointer;
         L     #TMP_dPZD_Pointer;
         +     16;
         T     #TMP_dPZD_Pointer;

         L     IW[ #TMP_dIO_Pointer];
         T     DIW[ #TMP_dPZD_Pointer];
END_REGION

REGION Network 6 (STL): Input copy power module
         L     #STC_tSYS_DATA.iIOAddress_PM;
         L     0;
         <=I;
         JC    NRPM;

         L     #STC_tSYS_DATA.iIOAddress_PM;
         SLW   3;
         T     #TMP_dIO_Pointer;

         L;
         T     #TMP_dPZD_Pointer;

         L     IW[ #TMP_dIO_Pointer];
         T     DIW[ #TMP_dPZD_Pointer];

         L     #STC_tSYS_DATA.iPowerOFFDelay_ms;
         L     1000;
         <I;
         JC    NWPM;

   NRPM: NOP   0;
END_REGION

REGION Network 7: Status signals